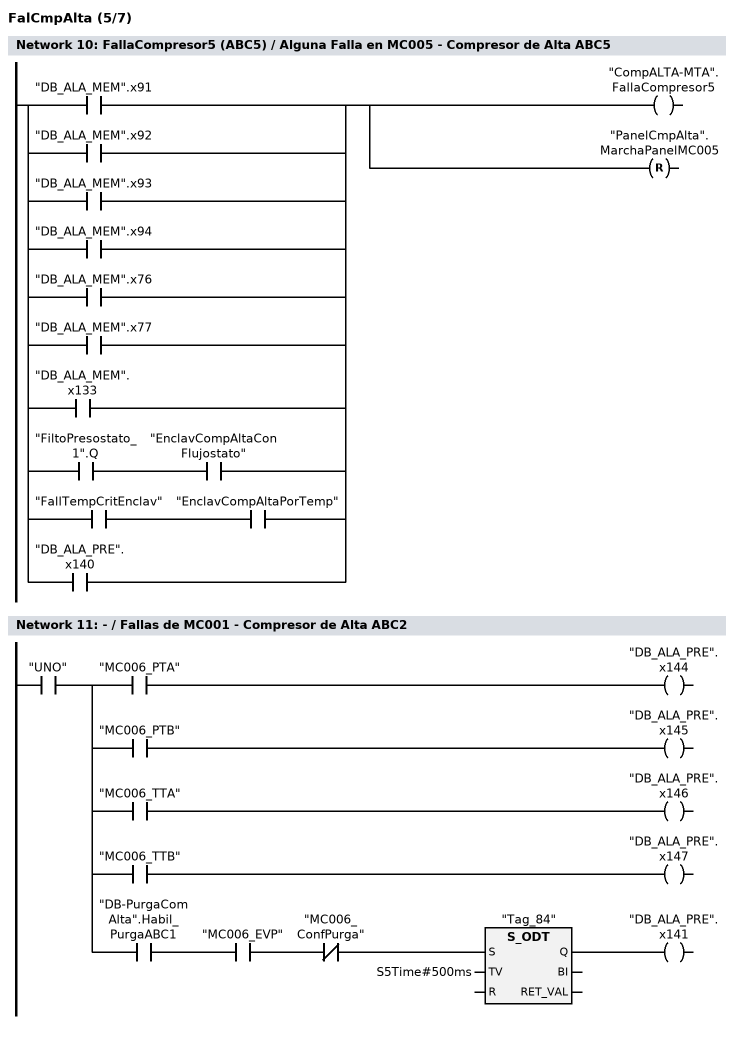
   RUNG wire#powerrail
      Contact( "DB_ALA_MEM".x91 )
      wire#w1
      Coil( "CompALTA-MTA".FallaCompresor5 )
   END_RUNG
   RUNG wire#powerrail
      Contact( "DB_ALA_MEM".x92 )
   END_RUNG wire#w1
   RUNG wire#powerrail
      Contact( "DB_ALA_MEM".x93 )
   END_RUNG wire#w1
   RUNG wire#powerrail
      Contact( "DB_ALA_MEM".x94 )
   END_RUNG wire#w1
   RUNG wire#powerrail
      Contact( "DB_ALA_MEM".x76 )
   END_RUNG wire#w1
   RUNG wire#powerrail
      Contact( "DB_ALA_MEM".x77 )
   END_RUNG wire#w1
   RUNG wire#powerrail
      Contact( "DB_ALA_MEM".x133 )
   END_RUNG wire#w1
   RUNG wire#powerrail
      Contact( "FiltoPresostato_1".Q )
      Contact( "EnclavCompAltaConFlujostato" )
   END_RUNG wire#w1
   RUNG wire#powerrail
      Contact( "FallTempCritEnclav" )
      Contact( "EnclavCompAltaPorTemp" )
   END_RUNG wire#w1
   RUNG wire#powerrail
      Contact( "DB_ALA_PRE".x140 )
   END_RUNG wire#w1
   RUNG wire#w1
      R_Coil( "PanelCmpAlta".MarchaPanelMC005 )
   END_RUNG
   // the same network as SCL:
   "CompALTA-MTA".FallaCompresor5 := "DB_ALA_MEM".x91 OR "DB_ALA_MEM".x92 OR "DB_ALA_MEM".x93 OR "DB_ALA_MEM".x94 OR "DB_ALA_MEM".x76 OR "DB_ALA_MEM".x77 OR "DB_ALA_MEM".x133 OR ("FiltoPresostato_1".Q AND "EnclavCompAltaConFlujostato") OR ("FallTempCritEnclav" AND "EnclavCompAltaPorTemp") OR "DB_ALA_PRE".x140;
   IF "CompALTA-MTA".FallaCompresor5 THEN "PanelCmpAlta".MarchaPanelMC005 := FALSE; END_IF;
END_REGION

REGION Network 11: - / Fallas de MC001 - Compresor de Alta ABC2
   RUNG wire#powerrail
      Contact( "UNO" )
      wire#w1
      Contact( "MC006_PTA" )
      Coil( "DB_ALA_PRE".x144 )
   END_RUNG
   RUNG wire#w1
      Contact( "MC006_PTB" )
      Coil( "DB_ALA_PRE".x145 )
   END_RUNG
   RUNG wire#w1
      Contact( "MC006_TTA" )
      Coil( "DB_ALA_PRE".x146 )
   END_RUNG
   RUNG wire#w1
      Contact( "MC006_TTB" )
      Coil( "DB_ALA_PRE".x147 )
   END_RUNG
   RUNG wire#w1
      Contact( "DB-PurgaComAlta".Habil_PurgaABC1 )
      Contact( "MC006_EVP" )
      I_Contact( "MC006_ConfPurga" )
      S_ODT(T_NO := "Tag_84", TV := S5Time#500ms, R :=, BI =>, RET_VAL =>)
      Coil( "DB_ALA_PRE".x141 )
   END_RUNG
   // the same network as SCL:
   "DB_ALA_PRE".x144 := "UNO" AND "MC006_PTA";
   "DB_ALA_PRE".x145 := "UNO" AND "MC006_PTB";
   "DB_ALA_PRE".x146 := "UNO" AND "MC006_TTA";
   "DB_ALA_PRE".x147 := "UNO" AND "MC006_TTB";
   #_s5time1 := S_ODT(T_NO := "Tag_84",
                      S := "UNO" AND "DB-PurgaComAlta".Habil_PurgaABC1 AND "MC006_EVP" AND NOT "MC006_ConfPurga",
                      TV := S5Time#500ms,
                      Q => #_w1);
   "DB_ALA_PRE".x141 := #_w1;
END_REGION

REGION Network 12: FallaCompresor6 (ABC1) / Alguna Falla en MC001 - Compresor de Alta ABC2
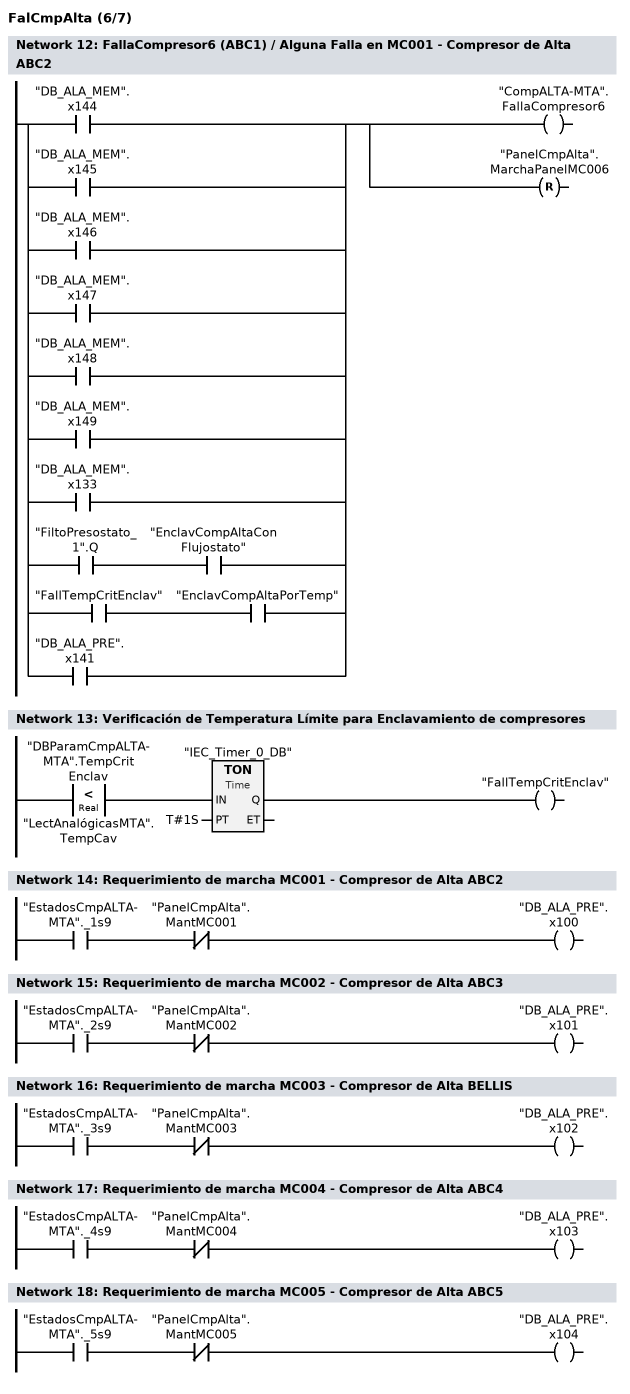
   RUNG wire#powerrail
      Contact( "DB_ALA_MEM".x144 )
      wire#w1
      Coil( "CompALTA-MTA".FallaCompresor6 )
   END_RUNG
   RUNG wire#powerrail
      Contact( "DB_ALA_MEM".x145 )
   END_RUNG wire#w1
   RUNG wire#powerrail
      Contact( "DB_ALA_MEM".x146 )
   END_RUNG wire#w1
   RUNG wire#powerrail
      Contact( "DB_ALA_MEM".x147 )
   END_RUNG wire#w1
   RUNG wire#powerrail
      Contact( "DB_ALA_MEM".x148 )
   END_RUNG wire#w1
   RUNG wire#powerrail
      Contact( "DB_ALA_MEM".x149 )
   END_RUNG wire#w1
   RUNG wire#powerrail
      Contact( "DB_ALA_MEM".x133 )
   END_RUNG wire#w1
   RUNG wire#powerrail
      Contact( "FiltoPresostato_1".Q )
      Contact( "EnclavCompAltaConFlujostato" )
   END_RUNG wire#w1
   RUNG wire#powerrail
      Contact( "FallTempCritEnclav" )
      Contact( "EnclavCompAltaPorTemp" )
   END_RUNG wire#w1
   RUNG wire#powerrail
      Contact( "DB_ALA_PRE".x141 )
   END_RUNG wire#w1
   RUNG wire#w1
      R_Coil( "PanelCmpAlta".MarchaPanelMC006 )
   END_RUNG
   // the same network as SCL:
   "CompALTA-MTA".FallaCompresor6 := "DB_ALA_MEM".x144 OR "DB_ALA_MEM".x145 OR "DB_ALA_MEM".x146 OR "DB_ALA_MEM".x147 OR "DB_ALA_MEM".x148 OR "DB_ALA_MEM".x149 OR "DB_ALA_MEM".x133 OR ("FiltoPresostato_1".Q AND "EnclavCompAltaConFlujostato") OR ("FallTempCritEnclav" AND "EnclavCompAltaPorTemp") OR "DB_ALA_PRE".x141;
   IF "CompALTA-MTA".FallaCompresor6 THEN "PanelCmpAlta".MarchaPanelMC006 := FALSE; END_IF;
END_REGION

REGION Network 13: Verificación de Temperatura Límite para Enclavamiento de compresores
   "IEC_Timer_0_DB".TON(IN := "DBParamCmpALTA-MTA".TempCritEnclav < "LectAnalógicasMTA".TempCav, PT := T#1S);
   "FallTempCritEnclav" := "IEC_Timer_0_DB".Q;
END_REGION

REGION Network 14: Requerimiento de marcha MC001 - Compresor de Alta ABC2
   RUNG wire#powerrail
      Contact( "EstadosCmpALTA-MTA"._1s9 )
      I_Contact( "PanelCmpAlta".MantMC001 )
      Coil( "DB_ALA_PRE".x100 )
   END_RUNG
   // the same network as SCL:
   "DB_ALA_PRE".x100 := "EstadosCmpALTA-MTA"._1s9 AND NOT "PanelCmpAlta".MantMC001;
END_REGION

REGION Network 15: Requerimiento de marcha MC002 - Compresor de Alta ABC3
   RUNG wire#powerrail
      Contact( "EstadosCmpALTA-MTA"._2s9 )
      I_Contact( "PanelCmpAlta".MantMC002 )
      Coil( "DB_ALA_PRE".x101 )
   END_RUNG
   // the same network as SCL:
   "DB_ALA_PRE".x101 := "EstadosCmpALTA-MTA"._2s9 AND NOT "PanelCmpAlta".MantMC002;
END_REGION

REGION Network 16: Requerimiento de marcha MC003 - Compresor de Alta BELLIS
   RUNG wire#powerrail
      Contact( "EstadosCmpALTA-MTA"._3s9 )
      I_Contact( "PanelCmpAlta".MantMC003 )
      Coil( "DB_ALA_PRE".x102 )
   END_RUNG
   // the same network as SCL:
   "DB_ALA_PRE".x102 := "EstadosCmpALTA-MTA"._3s9 AND NOT "PanelCmpAlta".MantMC003;
END_REGION

REGION Network 17: Requerimiento de marcha MC004 - Compresor de Alta ABC4
   RUNG wire#powerrail
      Contact( "EstadosCmpALTA-MTA"._4s9 )
      I_Contact( "PanelCmpAlta".MantMC004 )
      Coil( "DB_ALA_PRE".x103 )
   END_RUNG
   // the same network as SCL:
   "DB_ALA_PRE".x103 := "EstadosCmpALTA-MTA"._4s9 AND NOT "PanelCmpAlta".MantMC004;
END_REGION

REGION Network 18: Requerimiento de marcha MC005 - Compresor de Alta ABC5
   RUNG wire#powerrail
      Contact( "EstadosCmpALTA-MTA"._5s9 )
      I_Contact( "PanelCmpAlta".MantMC005 )
      Coil( "DB_ALA_PRE".x104 )
   END_RUNG
   // the same network as SCL:
   "DB_ALA_PRE".x104 := "EstadosCmpALTA-MTA"._5s9 AND NOT "PanelCmpAlta".MantMC005;
END_REGION

REGION Network 19: Requerimiento de marcha MC001 - Compresor de Alta ABC2
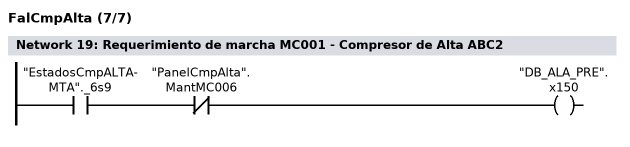
   RUNG wire#powerrail
      Contact( "EstadosCmpALTA-MTA"._6s9 )
      I_Contact( "PanelCmpAlta".MantMC006 )
      Coil( "DB_ALA_PRE".x150 )
   END_RUNG
   // the same network as SCL:
   "DB_ALA_PRE".x150 := "EstadosCmpALTA-MTA"._6s9 AND NOT "PanelCmpAlta".MantMC006;
END_REGION
END_FUNCTION

// folder: Auxiliares

FUNCTION "AjusteEntrada-SalidaMTA" : Void   // FC6, LAD
{ S7_Optimized_Access := 'FALSE' }
VERSION : 0.1
BEGIN

REGION Network 1
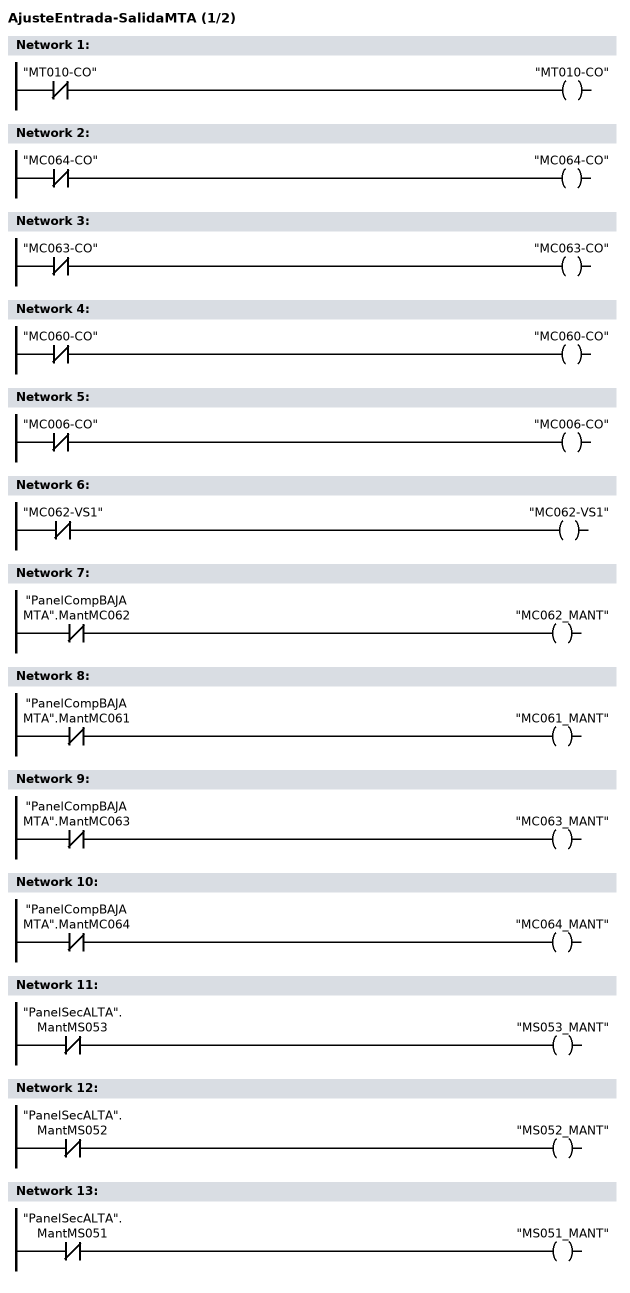
   RUNG wire#powerrail
      I_Contact( "MT010-CO" )
      Coil( "MT010-CO" )
   END_RUNG
   // the same network as SCL:
   "MT010-CO" := NOT "MT010-CO";
END_REGION

REGION Network 2
   RUNG wire#powerrail
      I_Contact( "MC064-CO" )
      Coil( "MC064-CO" )
   END_RUNG
   // the same network as SCL:
   "MC064-CO" := NOT "MC064-CO";
END_REGION

REGION Network 3
   RUNG wire#powerrail
      I_Contact( "MC063-CO" )
      Coil( "MC063-CO" )
   END_RUNG
   // the same network as SCL:
   "MC063-CO" := NOT "MC063-CO";
END_REGION

REGION Network 4
   RUNG wire#powerrail
      I_Contact( "MC060-CO" )
      Coil( "MC060-CO" )
   END_RUNG
   // the same network as SCL:
   "MC060-CO" := NOT "MC060-CO";
END_REGION

REGION Network 5
   RUNG wire#powerrail
      I_Contact( "MC006-CO" )
      Coil( "MC006-CO" )
   END_RUNG
   // the same network as SCL:
   "MC006-CO" := NOT "MC006-CO";
END_REGION

REGION Network 6
   RUNG wire#powerrail
      I_Contact( "MC062-VS1" )
      Coil( "MC062-VS1" )
   END_RUNG
   // the same network as SCL:
   "MC062-VS1" := NOT "MC062-VS1";
END_REGION

REGION Network 7
   RUNG wire#powerrail
      I_Contact( "PanelCompBAJA MTA".MantMC062 )
      Coil( "MC062_MANT" )
   END_RUNG
   // the same network as SCL:
   "MC062_MANT" := NOT "PanelCompBAJA MTA".MantMC062;
END_REGION

REGION Network 8
   RUNG wire#powerrail
      I_Contact( "PanelCompBAJA MTA".MantMC061 )
      Coil( "MC061_MANT" )
   END_RUNG
   // the same network as SCL:
   "MC061_MANT" := NOT "PanelCompBAJA MTA".MantMC061;
END_REGION

REGION Network 9
   RUNG wire#powerrail
      I_Contact( "PanelCompBAJA MTA".MantMC063 )
      Coil( "MC063_MANT" )
   END_RUNG
   // the same network as SCL:
   "MC063_MANT" := NOT "PanelCompBAJA MTA".MantMC063;
END_REGION

REGION Network 10
   RUNG wire#powerrail
      I_Contact( "PanelCompBAJA MTA".MantMC064 )
      Coil( "MC064_MANT" )
   END_RUNG
   // the same network as SCL:
   "MC064_MANT" := NOT "PanelCompBAJA MTA".MantMC064;
END_REGION

REGION Network 11
   RUNG wire#powerrail
      I_Contact( "PanelSecALTA".MantMS053 )
      Coil( "MS053_MANT" )
   END_RUNG
   // the same network as SCL:
   "MS053_MANT" := NOT "PanelSecALTA".MantMS053;
END_REGION

REGION Network 12
   RUNG wire#powerrail
      I_Contact( "PanelSecALTA".MantMS052 )
      Coil( "MS052_MANT" )
   END_RUNG
   // the same network as SCL:
   "MS052_MANT" := NOT "PanelSecALTA".MantMS052;
END_REGION

REGION Network 13
   RUNG wire#powerrail
      I_Contact( "PanelSecALTA".MantMS051 )
      Coil( "MS051_MANT" )
   END_RUNG
   // the same network as SCL:
   "MS051_MANT" := NOT "PanelSecALTA".MantMS051;
END_REGION

REGION Network 14
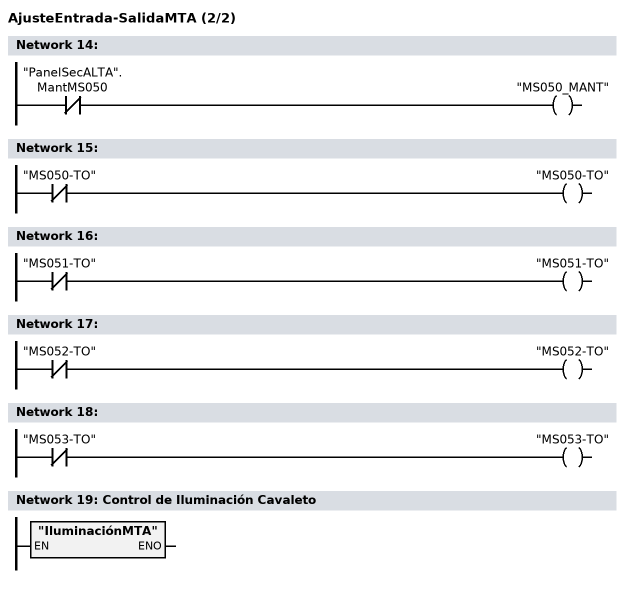
   RUNG wire#powerrail
      I_Contact( "PanelSecALTA".MantMS050 )
      Coil( "MS050_MANT" )
   END_RUNG
   // the same network as SCL:
   "MS050_MANT" := NOT "PanelSecALTA".MantMS050;
END_REGION

REGION Network 15
   RUNG wire#powerrail
      I_Contact( "MS050-TO" )
      Coil( "MS050-TO" )
   END_RUNG
   // the same network as SCL:
   "MS050-TO" := NOT "MS050-TO";
END_REGION

REGION Network 16
   RUNG wire#powerrail
      I_Contact( "MS051-TO" )
      Coil( "MS051-TO" )
   END_RUNG
   // the same network as SCL:
   "MS051-TO" := NOT "MS051-TO";
END_REGION

REGION Network 17
   RUNG wire#powerrail
      I_Contact( "MS052-TO" )
      Coil( "MS052-TO" )
   END_RUNG
   // the same network as SCL:
   "MS052-TO" := NOT "MS052-TO";
END_REGION

REGION Network 18
   RUNG wire#powerrail
      I_Contact( "MS053-TO" )
      Coil( "MS053-TO" )
   END_RUNG
   // the same network as SCL:
   "MS053-TO" := NOT "MS053-TO";
END_REGION

REGION Network 19: Control de Iluminación Cavaleto
   RUNG wire#powerrail
      "IluminaciónMTA"()
   END_RUNG
   // the same network as SCL:
   "IluminaciónMTA"();
END_REGION
END_FUNCTION

FUNCTION "And-Byte MTA" : Void   // FC22, LAD
{ S7_Optimized_Access := 'FALSE' }
VERSION : 0.1
BEGIN

REGION Network 1
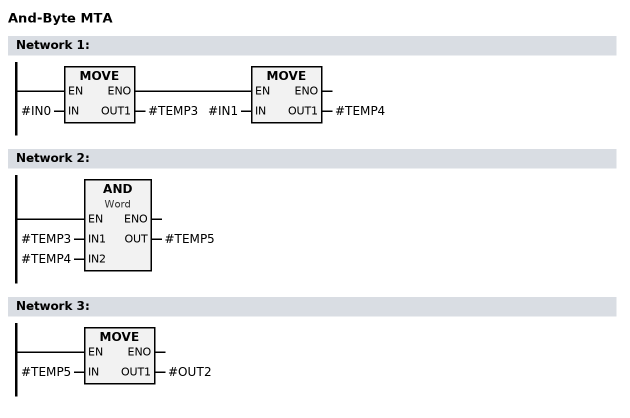
   RUNG wire#powerrail
      { S7_GenerateENO := "TRUE" } Move(in := #IN0, out1 => #TEMP3)
      { S7_GenerateENO := "TRUE" } Move(in := #IN1, out1 => #TEMP4)
   END_RUNG
   // the same network as SCL:
   // ENO of a box is taken as its EN; it also drops when the box reports an error
   #TEMP3 := #IN0;
   #TEMP4 := #IN1;
END_REGION

REGION Network 2
   RUNG wire#powerrail
      { S7_Templates := "SrcType := Word"; S7_GenerateENO := "TRUE" } And(in1 := #TEMP3, in2 := #TEMP4, out => #TEMP5)
   END_RUNG
   // the same network as SCL:
   #TEMP5 := #TEMP3 AND #TEMP4;
END_REGION

REGION Network 3
   RUNG wire#powerrail
      { S7_GenerateENO := "TRUE" } Move(in := #TEMP5, out1 => #OUT2)
   END_RUNG
   // the same network as SCL:
   #OUT2 := #TEMP5;
END_REGION
END_FUNCTION

FUNCTION "Inicialización" : Void   // FC46, LAD
{ S7_Optimized_Access := 'FALSE' }
VERSION : 0.1
BEGIN

REGION Network 1
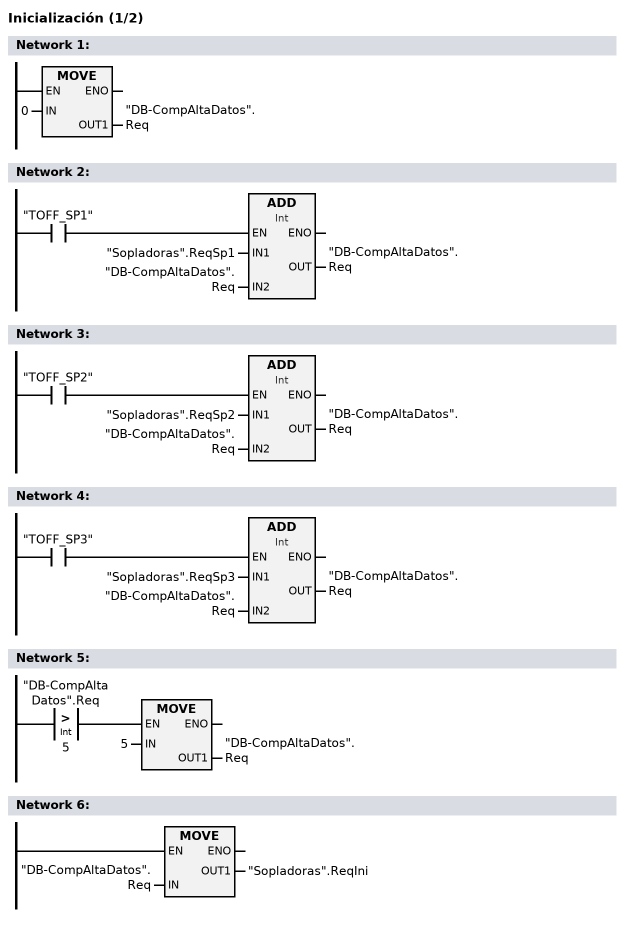
   RUNG wire#powerrail
      { S7_GenerateENO := "TRUE" } Move(in := 0, out1 => "DB-CompAltaDatos".Req)
   END_RUNG
   // the same network as SCL:
   "DB-CompAltaDatos".Req := 0;
END_REGION

REGION Network 2
   RUNG wire#powerrail
      Contact( "TOFF_SP1" )
      { S7_Templates := "SrcType := Int"; S7_GenerateENO := "TRUE" } Add(in1 := "Sopladoras".ReqSp1, in2 := "DB-CompAltaDatos".Req, out => "DB-CompAltaDatos".Req)
   END_RUNG
   // the same network as SCL:
   IF "TOFF_SP1" THEN "DB-CompAltaDatos".Req := "Sopladoras".ReqSp1 + "DB-CompAltaDatos".Req; END_IF;
END_REGION

REGION Network 3
   RUNG wire#powerrail
      Contact( "TOFF_SP2" )
      { S7_Templates := "SrcType := Int"; S7_GenerateENO := "TRUE" } Add(in1 := "Sopladoras".ReqSp2, in2 := "DB-CompAltaDatos".Req, out => "DB-CompAltaDatos".Req)
   END_RUNG
   // the same network as SCL:
   IF "TOFF_SP2" THEN "DB-CompAltaDatos".Req := "Sopladoras".ReqSp2 + "DB-CompAltaDatos".Req; END_IF;
END_REGION

REGION Network 4
   RUNG wire#powerrail
      Contact( "TOFF_SP3" )
      { S7_Templates := "SrcType := Int"; S7_GenerateENO := "TRUE" } Add(in1 := "Sopladoras".ReqSp3, in2 := "DB-CompAltaDatos".Req, out => "DB-CompAltaDatos".Req)
   END_RUNG
   // the same network as SCL:
   IF "TOFF_SP3" THEN "DB-CompAltaDatos".Req := "Sopladoras".ReqSp3 + "DB-CompAltaDatos".Req; END_IF;
END_REGION

REGION Network 5
   RUNG wire#powerrail
      { S7_Templates := "SrcType := Int" } GT_Contact(in1 := "DB-CompAltaDatos".Req, in2 := 5)
      { S7_GenerateENO := "TRUE" } Move(in := 5, out1 => "DB-CompAltaDatos".Req)
   END_RUNG
   // the same network as SCL:
   IF "DB-CompAltaDatos".Req > 5 THEN "DB-CompAltaDatos".Req := 5; END_IF;
END_REGION

REGION Network 6
   RUNG wire#powerrail
      { S7_GenerateENO := "TRUE" } Move(in := "DB-CompAltaDatos".Req, out1 => "Sopladoras".ReqIni)
   END_RUNG
   // the same network as SCL:
   "Sopladoras".ReqIni := "DB-CompAltaDatos".Req;
END_REGION

REGION Network 7
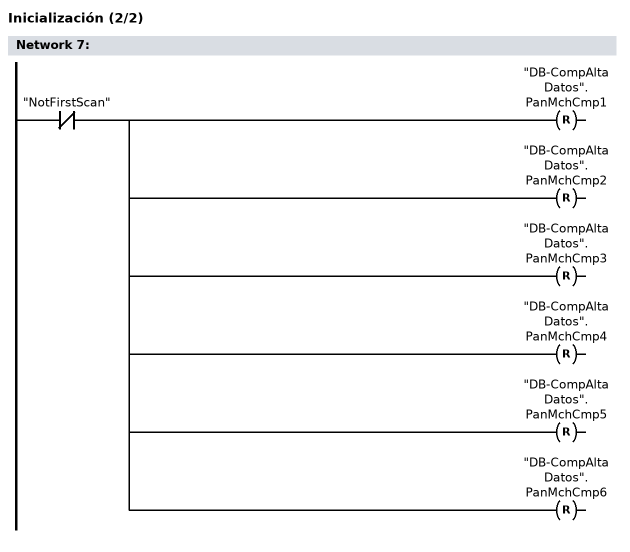
   RUNG wire#powerrail
      I_Contact( "NotFirstScan" )
      wire#w1
      R_Coil( "DB-CompAltaDatos".PanMchCmp1 )
   END_RUNG
   RUNG wire#w1
      R_Coil( "DB-CompAltaDatos".PanMchCmp2 )
   END_RUNG
   RUNG wire#w1
      R_Coil( "DB-CompAltaDatos".PanMchCmp3 )
   END_RUNG
   RUNG wire#w1
      R_Coil( "DB-CompAltaDatos".PanMchCmp4 )
   END_RUNG
   RUNG wire#w1
      R_Coil( "DB-CompAltaDatos".PanMchCmp5 )
   END_RUNG
   RUNG wire#w1
      R_Coil( "DB-CompAltaDatos".PanMchCmp6 )
   END_RUNG
   // the same network as SCL:
   IF NOT "NotFirstScan" THEN
       "DB-CompAltaDatos".PanMchCmp1 := FALSE;
       "DB-CompAltaDatos".PanMchCmp2 := FALSE;
       "DB-CompAltaDatos".PanMchCmp3 := FALSE;
       "DB-CompAltaDatos".PanMchCmp4 := FALSE;
       "DB-CompAltaDatos".PanMchCmp5 := FALSE;
       "DB-CompAltaDatos".PanMchCmp6 := FALSE;
   END_IF;
END_REGION
END_FUNCTION

// folder: Bloques Estándar

FUNCTION_BLOCK "ControladorMotoresMTA"   // FB2, LAD
{ S7_Optimized_Access := 'FALSE' }
VERSION : 0.1
BEGIN

REGION Network 2
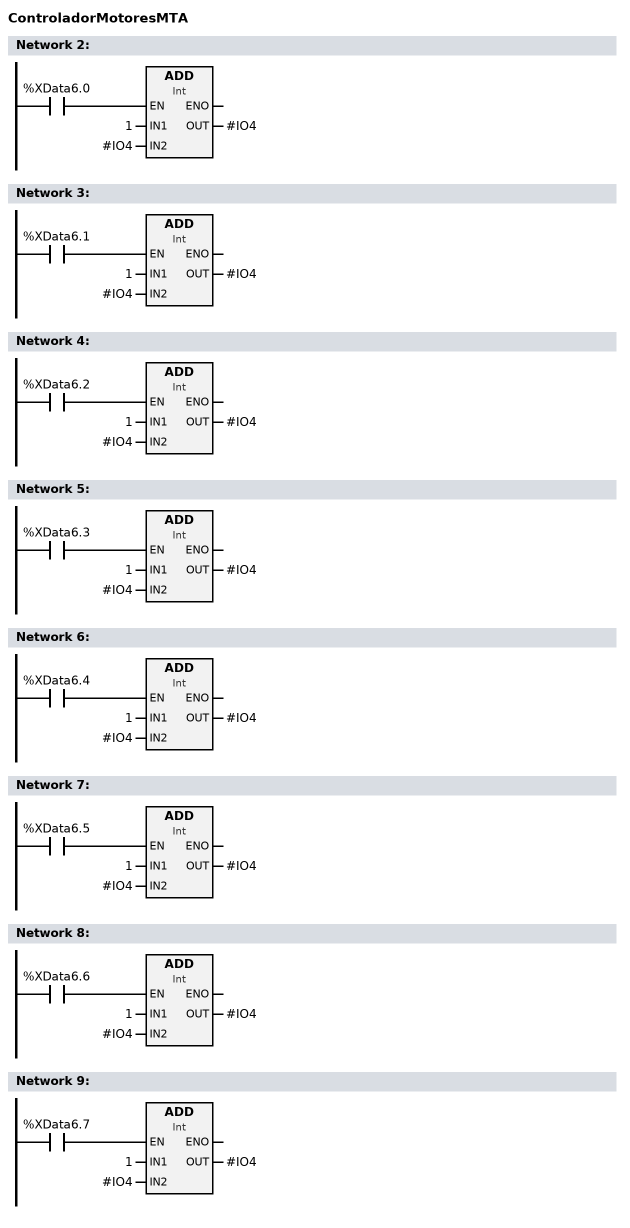
   RUNG wire#powerrail
      Contact( %XData6.0 )
      { S7_Templates := "SrcType := Int"; S7_GenerateENO := "TRUE" } Add(in1 := 1, in2 := #IO4, out => #IO4)
   END_RUNG
   // the same network as SCL:
   IF %XData6.0 THEN #IO4 := 1 + #IO4; END_IF;
END_REGION

REGION Network 3
   RUNG wire#powerrail
      Contact( %XData6.1 )
      { S7_Templates := "SrcType := Int"; S7_GenerateENO := "TRUE" } Add(in1 := 1, in2 := #IO4, out => #IO4)
   END_RUNG
   // the same network as SCL:
   IF %XData6.1 THEN #IO4 := 1 + #IO4; END_IF;
END_REGION

REGION Network 4
   RUNG wire#powerrail
      Contact( %XData6.2 )
      { S7_Templates := "SrcType := Int"; S7_GenerateENO := "TRUE" } Add(in1 := 1, in2 := #IO4, out => #IO4)
   END_RUNG
   // the same network as SCL:
   IF %XData6.2 THEN #IO4 := 1 + #IO4; END_IF;
END_REGION

REGION Network 5
   RUNG wire#powerrail
      Contact( %XData6.3 )
      { S7_Templates := "SrcType := Int"; S7_GenerateENO := "TRUE" } Add(in1 := 1, in2 := #IO4, out => #IO4)
   END_RUNG
   // the same network as SCL:
   IF %XData6.3 THEN #IO4 := 1 + #IO4; END_IF;
END_REGION

REGION Network 6
   RUNG wire#powerrail
      Contact( %XData6.4 )
      { S7_Templates := "SrcType := Int"; S7_GenerateENO := "TRUE" } Add(in1 := 1, in2 := #IO4, out => #IO4)
   END_RUNG
   // the same network as SCL:
   IF %XData6.4 THEN #IO4 := 1 + #IO4; END_IF;
END_REGION

REGION Network 7
   RUNG wire#powerrail
      Contact( %XData6.5 )
      { S7_Templates := "SrcType := Int"; S7_GenerateENO := "TRUE" } Add(in1 := 1, in2 := #IO4, out => #IO4)
   END_RUNG
   // the same network as SCL:
   IF %XData6.5 THEN #IO4 := 1 + #IO4; END_IF;
END_REGION

REGION Network 8
   RUNG wire#powerrail
      Contact( %XData6.6 )
      { S7_Templates := "SrcType := Int"; S7_GenerateENO := "TRUE" } Add(in1 := 1, in2 := #IO4, out => #IO4)
   END_RUNG
   // the same network as SCL:
   IF %XData6.6 THEN #IO4 := 1 + #IO4; END_IF;
END_REGION

REGION Network 9
   RUNG wire#powerrail
      Contact( %XData6.7 )
      { S7_Templates := "SrcType := Int"; S7_GenerateENO := "TRUE" } Add(in1 := 1, in2 := #IO4, out => #IO4)
   END_RUNG
   // the same network as SCL:
   IF %XData6.7 THEN #IO4 := 1 + #IO4; END_IF;
END_REGION
END_FUNCTION_BLOCK

// folder: Bloques Estándar/Boosters

FUNCTION "Booster (MTA)" : Void   // FC25, LAD
TITLE = Manejo General de los Boosters
{ S7_Optimized_Access := 'FALSE' }
VERSION : 0.1
   VAR_TEMP   // added for the SCL form of the ladder/FBD networks
      _w1 : Bool;
      _s5time1 : S5Time;
      _w2 : Bool;
      _s5time2 : S5Time;
      _w3 : Bool;
   END_VAR
BEGIN

REGION Network 1: Validación Horas para invertir prioridades
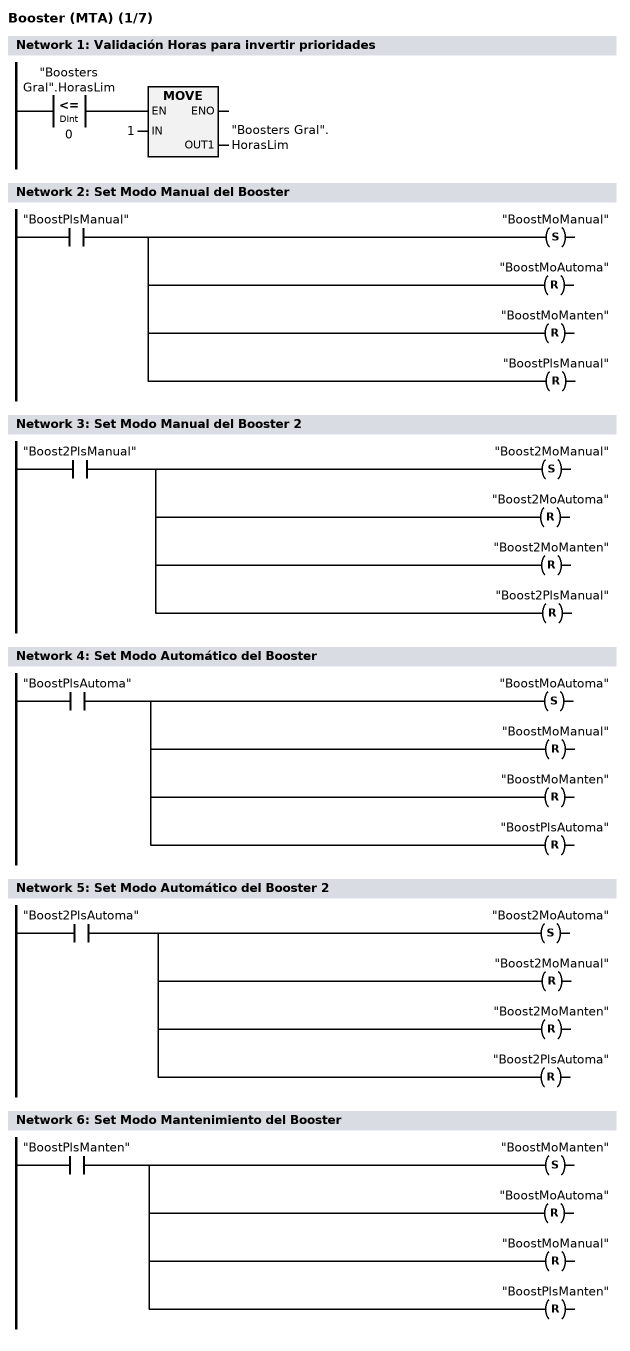
   RUNG wire#powerrail
      { S7_Templates := "SrcType := DInt" } LE_Contact(in1 := "Boosters Gral".HorasLim, in2 := 0)
      { S7_GenerateENO := "TRUE" } Move(in := 1, out1 => "Boosters Gral".HorasLim)
   END_RUNG
   // the same network as SCL:
   IF "Boosters Gral".HorasLim <= 0 THEN "Boosters Gral".HorasLim := 1; END_IF;
END_REGION

REGION Network 2: Set Modo Manual del Booster
   RUNG wire#powerrail
      Contact( "BoostPlsManual" )
      wire#w1
      S_Coil( "BoostMoManual" )
   END_RUNG
   RUNG wire#w1
      R_Coil( "BoostMoAutoma" )
   END_RUNG
   RUNG wire#w1
      R_Coil( "BoostMoManten" )
   END_RUNG
   RUNG wire#w1
      R_Coil( "BoostPlsManual" )
   END_RUNG
   // the same network as SCL:
   IF "BoostPlsManual" THEN
       "BoostMoManual" := TRUE;
       "BoostMoAutoma" := FALSE;
       "BoostMoManten" := FALSE;
       "BoostPlsManual" := FALSE;
   END_IF;
END_REGION

REGION Network 3: Set Modo Manual del Booster 2
   RUNG wire#powerrail
      Contact( "Boost2PlsManual" )
      wire#w1
      S_Coil( "Boost2MoManual" )
   END_RUNG
   RUNG wire#w1
      R_Coil( "Boost2MoAutoma" )
   END_RUNG
   RUNG wire#w1
      R_Coil( "Boost2MoManten" )
   END_RUNG
   RUNG wire#w1
      R_Coil( "Boost2PlsManual" )
   END_RUNG
   // the same network as SCL:
   IF "Boost2PlsManual" THEN
       "Boost2MoManual" := TRUE;
       "Boost2MoAutoma" := FALSE;
       "Boost2MoManten" := FALSE;
       "Boost2PlsManual" := FALSE;
   END_IF;
END_REGION

REGION Network 4: Set Modo Automático del Booster
   RUNG wire#powerrail
      Contact( "BoostPlsAutoma" )
      wire#w1
      S_Coil( "BoostMoAutoma" )
   END_RUNG
   RUNG wire#w1
      R_Coil( "BoostMoManual" )
   END_RUNG
   RUNG wire#w1
      R_Coil( "BoostMoManten" )
   END_RUNG
   RUNG wire#w1
      R_Coil( "BoostPlsAutoma" )
   END_RUNG
   // the same network as SCL:
   IF "BoostPlsAutoma" THEN
       "BoostMoAutoma" := TRUE;
       "BoostMoManual" := FALSE;
       "BoostMoManten" := FALSE;
       "BoostPlsAutoma" := FALSE;
   END_IF;
END_REGION

REGION Network 5: Set Modo Automático del Booster 2
   RUNG wire#powerrail
      Contact( "Boost2PlsAutoma" )
      wire#w1
      S_Coil( "Boost2MoAutoma" )
   END_RUNG
   RUNG wire#w1
      R_Coil( "Boost2MoManual" )
   END_RUNG
   RUNG wire#w1
      R_Coil( "Boost2MoManten" )
   END_RUNG
   RUNG wire#w1
      R_Coil( "Boost2PlsAutoma" )
   END_RUNG
   // the same network as SCL:
   IF "Boost2PlsAutoma" THEN
       "Boost2MoAutoma" := TRUE;
       "Boost2MoManual" := FALSE;
       "Boost2MoManten" := FALSE;
       "Boost2PlsAutoma" := FALSE;
   END_IF;
END_REGION

REGION Network 6: Set Modo Mantenimiento del Booster
   RUNG wire#powerrail
      Contact( "BoostPlsManten" )
      wire#w1
      S_Coil( "BoostMoManten" )
   END_RUNG
   RUNG wire#w1
      R_Coil( "BoostMoAutoma" )
   END_RUNG
   RUNG wire#w1
      R_Coil( "BoostMoManual" )
   END_RUNG
   RUNG wire#w1
      R_Coil( "BoostPlsManten" )
   END_RUNG
   // the same network as SCL:
   IF "BoostPlsManten" THEN
       "BoostMoManten" := TRUE;
       "BoostMoAutoma" := FALSE;
       "BoostMoManual" := FALSE;
       "BoostPlsManten" := FALSE;
   END_IF;
END_REGION

REGION Network 7: Set Modo Mantenimiento del Booster 2
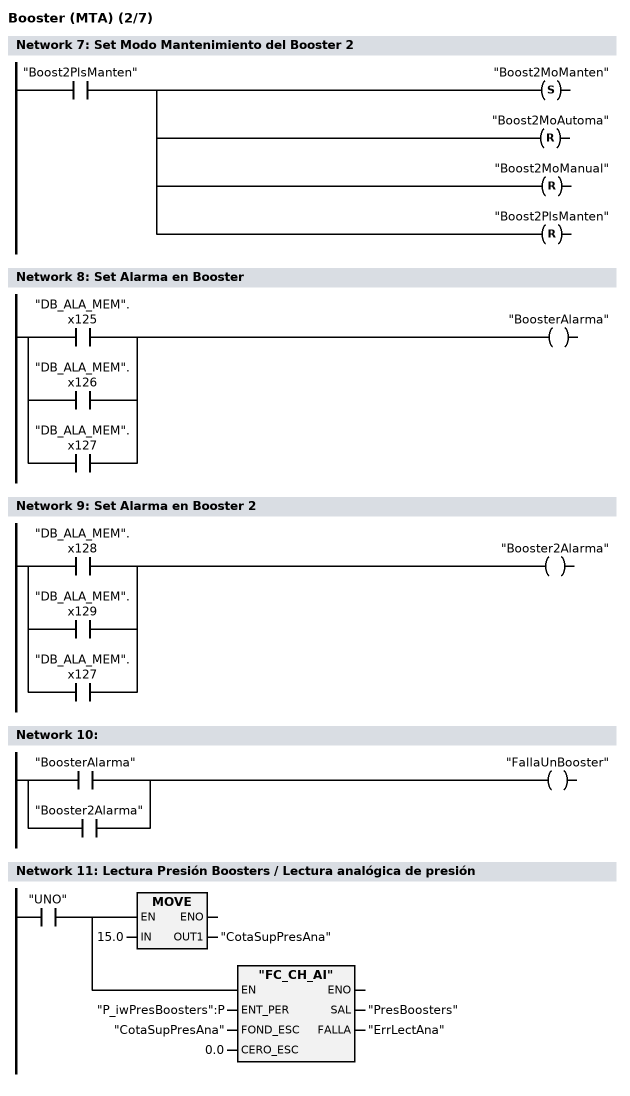
   RUNG wire#powerrail
      Contact( "Boost2PlsManten" )
      wire#w1
      S_Coil( "Boost2MoManten" )
   END_RUNG
   RUNG wire#w1
      R_Coil( "Boost2MoAutoma" )
   END_RUNG
   RUNG wire#w1
      R_Coil( "Boost2MoManual" )
   END_RUNG
   RUNG wire#w1
      R_Coil( "Boost2PlsManten" )
   END_RUNG
   // the same network as SCL:
   IF "Boost2PlsManten" THEN
       "Boost2MoManten" := TRUE;
       "Boost2MoAutoma" := FALSE;
       "Boost2MoManual" := FALSE;
       "Boost2PlsManten" := FALSE;
   END_IF;
END_REGION

REGION Network 8: Set Alarma en Booster
   RUNG wire#powerrail
      Contact( "DB_ALA_MEM".x125 )
      wire#w1
      Coil( "BoosterAlarma" )
   END_RUNG
   RUNG wire#powerrail
      Contact( "DB_ALA_MEM".x126 )
   END_RUNG wire#w1
   RUNG wire#powerrail
      Contact( "DB_ALA_MEM".x127 )
   END_RUNG wire#w1
   // the same network as SCL:
   "BoosterAlarma" := "DB_ALA_MEM".x125 OR "DB_ALA_MEM".x126 OR "DB_ALA_MEM".x127;
END_REGION

REGION Network 9: Set Alarma en Booster 2
   RUNG wire#powerrail
      Contact( "DB_ALA_MEM".x128 )
      wire#w1
      Coil( "Booster2Alarma" )
   END_RUNG
   RUNG wire#powerrail
      Contact( "DB_ALA_MEM".x129 )
   END_RUNG wire#w1
   RUNG wire#powerrail
      Contact( "DB_ALA_MEM".x127 )
   END_RUNG wire#w1
   // the same network as SCL:
   "Booster2Alarma" := "DB_ALA_MEM".x128 OR "DB_ALA_MEM".x129 OR "DB_ALA_MEM".x127;
END_REGION

REGION Network 10
   RUNG wire#powerrail
      Contact( "BoosterAlarma" )
      wire#w1
      Coil( "FallaUnBooster" )
   END_RUNG
   RUNG wire#powerrail
      Contact( "Booster2Alarma" )
   END_RUNG wire#w1
   // the same network as SCL:
   "FallaUnBooster" := "BoosterAlarma" OR "Booster2Alarma";
END_REGION

REGION Network 11: Lectura Presión Boosters / Lectura analógica de presión
   RUNG wire#powerrail
      Contact( "UNO" )
      wire#w1
      { S7_GenerateENO := "TRUE" } Move(in := 15.0, out1 => "CotaSupPresAna")
   END_RUNG
   RUNG wire#w1
      "FC_CH_AI"(ENT_PER := "P_iwPresBoosters":P, FOND_ESC := "CotaSupPresAna", CERO_ESC := 0.0, SAL => "PresBoosters", FALLA => "ErrLectAna")
   END_RUNG
   // the same network as SCL:
   IF "UNO" THEN
       "CotaSupPresAna" := 15.0;
       "FC_CH_AI"(ENT_PER := "P_iwPresBoosters":P,
                  FOND_ESC := "CotaSupPresAna",
                  CERO_ESC := 0.0,
                  SAL => "PresBoosters",
                  FALLA => "ErrLectAna");
   END_IF;
END_REGION

REGION Network 12: Bandas de presión para arranque de Boosters / Set-Reset para control analógico
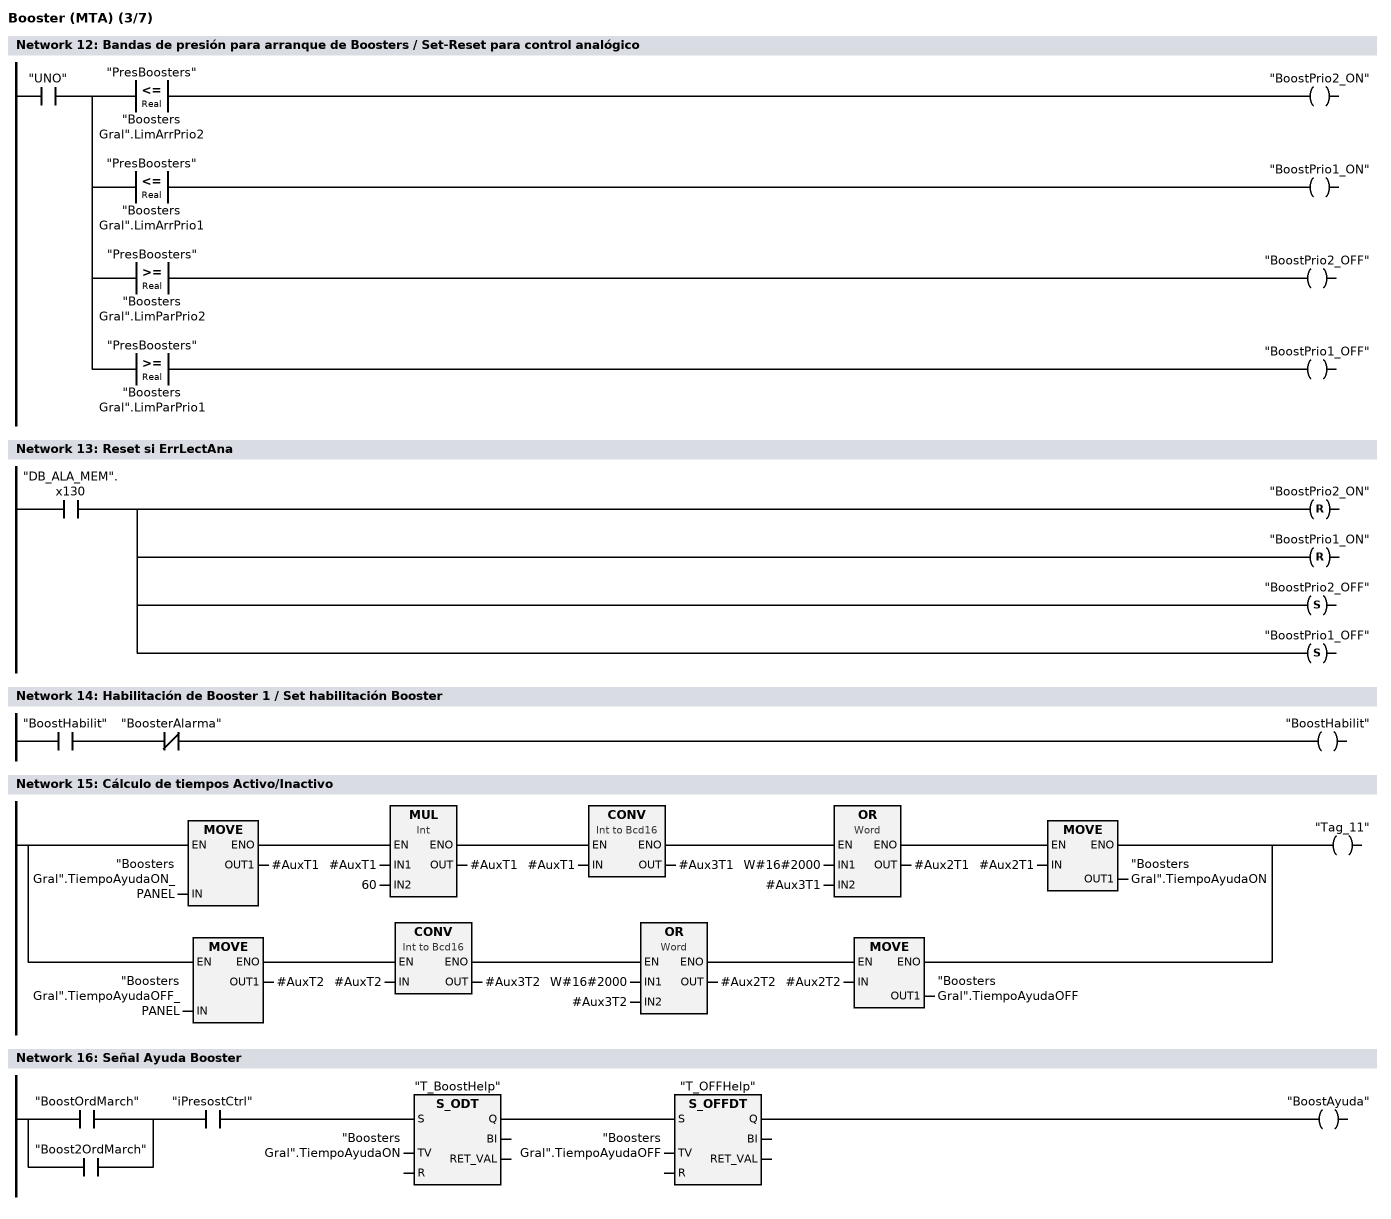
   RUNG wire#powerrail
      Contact( "UNO" )
      wire#w1
      { S7_Templates := "SrcType := Real" } LE_Contact(in1 := "PresBoosters", in2 := "Boosters Gral".LimArrPrio2)
      Coil( "BoostPrio2_ON" )
   END_RUNG
   RUNG wire#w1
      { S7_Templates := "SrcType := Real" } LE_Contact(in1 := "PresBoosters", in2 := "Boosters Gral".LimArrPrio1)
      Coil( "BoostPrio1_ON" )
   END_RUNG
   RUNG wire#w1
      { S7_Templates := "SrcType := Real" } GE_Contact(in1 := "PresBoosters", in2 := "Boosters Gral".LimParPrio2)
      Coil( "BoostPrio2_OFF" )
   END_RUNG
   RUNG wire#w1
      { S7_Templates := "SrcType := Real" } GE_Contact(in1 := "PresBoosters", in2 := "Boosters Gral".LimParPrio1)
      Coil( "BoostPrio1_OFF" )
   END_RUNG
   // the same network as SCL:
   "BoostPrio2_ON" := "UNO" AND ("PresBoosters" <= "Boosters Gral".LimArrPrio2);
   "BoostPrio1_ON" := "UNO" AND ("PresBoosters" <= "Boosters Gral".LimArrPrio1);
   "BoostPrio2_OFF" := "UNO" AND ("PresBoosters" >= "Boosters Gral".LimParPrio2);
   "BoostPrio1_OFF" := "UNO" AND ("PresBoosters" >= "Boosters Gral".LimParPrio1);
END_REGION

REGION Network 13: Reset si ErrLectAna
   RUNG wire#powerrail
      Contact( "DB_ALA_MEM".x130 )
      wire#w1
      R_Coil( "BoostPrio2_ON" )
   END_RUNG
   RUNG wire#w1
      R_Coil( "BoostPrio1_ON" )
   END_RUNG
   RUNG wire#w1
      S_Coil( "BoostPrio2_OFF" )
   END_RUNG
   RUNG wire#w1
      S_Coil( "BoostPrio1_OFF" )
   END_RUNG
   // the same network as SCL:
   IF "DB_ALA_MEM".x130 THEN
       "BoostPrio2_ON" := FALSE;
       "BoostPrio1_ON" := FALSE;
       "BoostPrio2_OFF" := TRUE;
       "BoostPrio1_OFF" := TRUE;
   END_IF;
END_REGION

REGION Network 14: Habilitación de Booster 1 / Set habilitación Booster
   RUNG wire#powerrail
      Contact( "BoostHabilit" )
      I_Contact( "BoosterAlarma" )
      Coil( "BoostHabilit" )
   END_RUNG
   // the same network as SCL:
   "BoostHabilit" := "BoostHabilit" AND NOT "BoosterAlarma";
END_REGION

REGION Network 15: Cálculo de tiempos Activo/Inactivo
   // no checked SCL form for this network; see the picture
END_REGION

REGION Network 16: Señal Ayuda Booster
   RUNG wire#powerrail
      Contact( "BoostOrdMarch" )
      wire#w1
      Contact( "iPresostCtrl" )
      S_ODT(T_NO := "T_BoostHelp", TV := "Boosters Gral".TiempoAyudaON, R :=, BI =>, RET_VAL =>)
      S_OFFDT(T_NO := "T_OFFHelp", TV := "Boosters Gral".TiempoAyudaOFF, R :=, BI =>, RET_VAL =>)
      Coil( "BoostAyuda" )
   END_RUNG
   RUNG wire#powerrail
      Contact( "Boost2OrdMarch" )
   END_RUNG wire#w1
   // the same network as SCL:
   #_s5time1 := S_ODT(T_NO := "T_BoostHelp",
                      S := ("BoostOrdMarch" OR "Boost2OrdMarch") AND "iPresostCtrl",
                      TV := "Boosters Gral".TiempoAyudaON,
                      Q => #_w1);
   #_s5time2 := S_OFFDT(T_NO := "T_OFFHelp", S := #_w1, TV := "Boosters Gral".TiempoAyudaOFF, Q => #_w2);
   "BoostAyuda" := #_w2;
END_REGION

REGION Network 17: Prioridades Boosters / Prioridades Nulas
